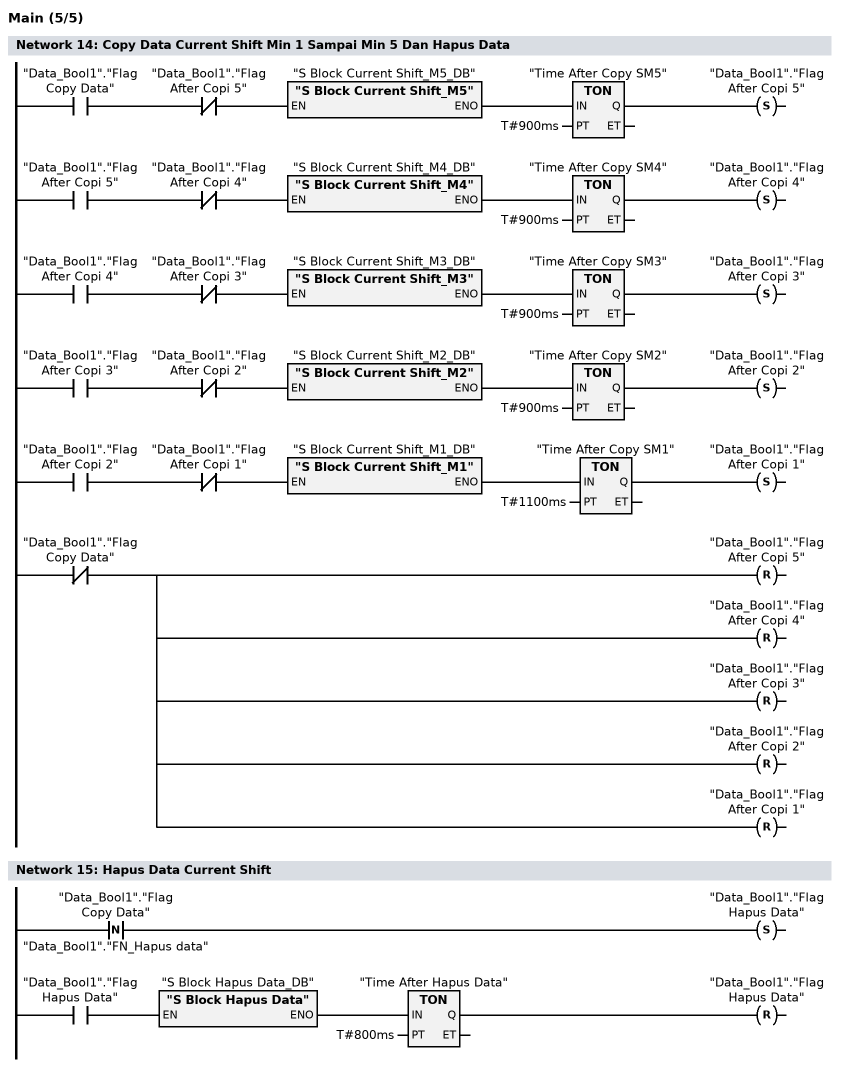
   "S Block Current Shift_M5_DB"(EN := "Data_Bool1"."Flag Copy Data" AND NOT "Data_Bool1"."Flag After Copi 5",   // "S Block Current Shift_M5"
                           ENO => #_w1);
   "Time After Copy SM5".TON(IN := #_w1, PT := T#900ms);
   IF "Time After Copy SM5".Q THEN "Data_Bool1"."Flag After Copi 5" := TRUE; END_IF;
   "S Block Current Shift_M4_DB"(EN := "Data_Bool1"."Flag After Copi 5" AND NOT "Data_Bool1"."Flag After Copi 4",   // "S Block Current Shift_M4"
                           ENO => #_w2);
   "Time After Copy SM4".TON(IN := #_w2, PT := T#900ms);
   IF "Time After Copy SM4".Q THEN "Data_Bool1"."Flag After Copi 4" := TRUE; END_IF;
   "S Block Current Shift_M3_DB"(EN := "Data_Bool1"."Flag After Copi 4" AND NOT "Data_Bool1"."Flag After Copi 3",   // "S Block Current Shift_M3"
                           ENO => #_w3);
   "Time After Copy SM3".TON(IN := #_w3, PT := T#900ms);
   IF "Time After Copy SM3".Q THEN "Data_Bool1"."Flag After Copi 3" := TRUE; END_IF;
   "S Block Current Shift_M2_DB"(EN := "Data_Bool1"."Flag After Copi 3" AND NOT "Data_Bool1"."Flag After Copi 2",   // "S Block Current Shift_M2"
                           ENO => #_w4);
   "Time After Copy SM2".TON(IN := #_w4, PT := T#900ms);
   IF "Time After Copy SM2".Q THEN "Data_Bool1"."Flag After Copi 2" := TRUE; END_IF;
   "S Block Current Shift_M1_DB"(EN := "Data_Bool1"."Flag After Copi 2" AND NOT "Data_Bool1"."Flag After Copi 1",   // "S Block Current Shift_M1"
                           ENO => #_w5);
   "Time After Copy SM1".TON(IN := #_w5, PT := T#1100ms);
   IF "Time After Copy SM1".Q THEN "Data_Bool1"."Flag After Copi 1" := TRUE; END_IF;
   IF NOT "Data_Bool1"."Flag Copy Data" THEN
       "Data_Bool1"."Flag After Copi 5" := FALSE;
       "Data_Bool1"."Flag After Copi 4" := FALSE;
       "Data_Bool1"."Flag After Copi 3" := FALSE;
       "Data_Bool1"."Flag After Copi 2" := FALSE;
       "Data_Bool1"."Flag After Copi 1" := FALSE;
   END_IF;
END_REGION

REGION Network 15: Hapus Data Current Shift
   #_w1 := NOT "Data_Bool1"."Flag Copy Data" AND "Data_Bool1"."FN_Hapus data";   // falling edge of "Data_Bool1"."Flag Copy Data"
   "Data_Bool1"."FN_Hapus data" := "Data_Bool1"."Flag Copy Data";
   IF #_w1 THEN "Data_Bool1"."Flag Hapus Data" := TRUE; END_IF;
   "S Block Hapus Data_DB"(EN := "Data_Bool1"."Flag Hapus Data", ENO => #_w2);   // "S Block Hapus Data"
   "Time After Hapus Data".TON(IN := #_w2, PT := T#800ms);
   IF "Time After Hapus Data".Q THEN "Data_Bool1"."Flag Hapus Data" := FALSE; END_IF;
END_REGION
END_ORGANIZATION_BLOCK

ORGANIZATION_BLOCK "Time error interrupt"   // OB80, LAD, TimeErrorInterrupt
{ S7_Optimized_Access := 'TRUE' }
VERSION : 0.1
   VAR_INPUT
      Fault_ID : Byte;   // Fault identifier
      Csg_OBnr : OB_Any;   // Number of OB causing the error
      Csg_Prio : UInt;   // Priority of OB causing the error
   END_VAR
BEGIN
END_ORGANIZATION_BLOCK

ORGANIZATION_BLOCK "Diagnostic error interrupt"   // OB82, LAD, DiagnosticErrorInterrupt
{ S7_Optimized_Access := 'TRUE' }
VERSION : 0.1
   VAR_INPUT
      IO_State : Word;   // IO state of the HW object
      LADDR : Hw_Any;   // Hardware identifier
      Channel : UInt;   // Channel number
      MultiError : Bool;   // =true if more than one error is present
   END_VAR
BEGIN
END_ORGANIZATION_BLOCK

(* ===== HMI "HMI_RT_1" =====
system functions are stored by id; their names below are inferred from use
connection "HMI_connection": ETHERNET, SMART_S7_1200_OMS

HMI tags "Default tag table"
   "Tag_ScreenNumber" : UInt, internal
      on ChangeValue: ActivateScreenByNumber("Tag_ScreenNumber", 0)
   "PB Test Pneumatic 1" : Bool = PLC "PB Test Pneumatic 1" AT %M205.1, 1 s
   "PB Test Pneumatic 2" : Bool = PLC "PB Test Pneumatic 2" AT %M205.2, 1 s
   "PB Test Pneumatic 3" : Bool = PLC "PB Test Pneumatic 3" AT %M205.3, 1 s
   "PB Test Pneumatic 4" : Bool = PLC "PB Test Pneumatic 4" AT %M205.4, 1 s
   "PB Test Pneumatic 5" : Bool = PLC "PB Test Pneumatic 5" AT %M205.5, 1 s
   "PB Test Motor" : Bool = PLC "PB Test Motor" AT %M205.7, 1 s
   "PB Test Manual Servo" : Bool = PLC "PB Test Manual Servo" AT %M205.6, 1 s
   "Timer Waktu Pemanasan" : Time = PLC "Timer Delay Heating" AT %MD0, 1 s
   "Machine Running" : Bool = PLC "Machine Running" AT %M200.0, 1 s
   "Flag Imaje Start" : Bool = PLC "Flag Imaje Start" AT %M212.0, 1 s
   "Counter" : Int = PLC Counter AT %MW5, 1 s
   "Counter Ejector" : Int = PLC "Counter Ejector" AT %MW9, 1 s
   "Reset Counter" : Bool = PLC "Reset Counter" AT %M200.1, 1 s
   "PB Test Mode" : Bool = PLC "PB Test Mode" AT %M205.0, 1 s
   "Flag Ejector Jalan" : Bool = PLC "Flag Ejector Jalan" AT %M230.3, 1 s
   "Error Group" : Word = PLC "Error Group" AT %MW4, 1 s
   "PB Test Imaje" : Bool = PLC "PB Test Imaje" AT %M206.0, 1 s
   "PB Test Air Valve" : Bool = PLC "PB Test Air Valve" AT %M206.1, 1 s
   "Flag Barcode HMI" : Bool = PLC "Flag Enable/Disable Barcode HMI" AT %M30.0, 1 s
   "Flag Enable/Disable Error Chute 3 Way" : Bool = PLC "Flag Enable/Disable Error Chute 3 Way" AT %M30.1, 1 s
   "Flag Parameter Page" : Bool = PLC "Flag Parameter Page" AT %M232.6, 1 s
   "Flag Main Page" : Bool = PLC "Flag Main Page" AT %M232.7, 1 s
   "HMI_Tag_1" : Word AT %DB39.DBW0, 1 s
   "HMI_Error_Cont" : Word AT %DB40.DBW0, 1 s
   "Flag Teach In Barcode" : Bool = PLC "Flag Teach In Barcode" AT %M212.4, 1 s
   "Teach In Barcode" : Bool = PLC "Teach In Barcode" AT %Q0.5, 1 s
   "Flag Heater Error HMI" : Bool = PLC "Flag Heater Error HMI" AT %M30.2, 1 s
   "Flag Pneumatic Bypass" : Bool = PLC "Flag Reed Switch Bypass" AT %M30.3, 1 s
   "Flag Enable/Disable Error Door Open" : Bool = PLC "Flag Enable/Disable Error Door Open" AT %M30.5, 1 s
   "Timer Delay Stamp" : Time = PLC "Timer Delay Stamp" AT %MD32, 1 s
   "Flag Enable/Disable Block Focke" : Bool = PLC "Flag Enable/Disable Block Focke" AT %M30.6, 1 s
   "Flag Enable/Disable Error Chute Before Heating Roll" : Bool = PLC "Flag Enable/Disable Error Chute Before Heating Roll" AT %M30.4, 1 s
   "Flag Machine Bypass" : Bool = PLC "Flag Machine Bypass" AT %M30.7, 1 s
   "RS Bypass Pneumatic 1" : Bool = PLC "RS Bypass Pneumatic 1" AT %M31.0, 1 s
   "RS Bypass Pneumatic 3" : Bool = PLC "RS Bypass Pneumatic 3" AT %M31.1, 1 s
   "RS Bypass Pneumatic 4" : Bool = PLC "RS Bypass Pneumatic 4" AT %M31.2, 1 s
   "RS Bypass Pneumatic 5" : Bool = PLC "RS Bypass Pneumatic 5" AT %M31.3, 1 s
   "PB Test Pneumatic 6" : Bool = PLC "PB Test Pneumatic 6" AT %M206.2, 1 s
   "PB Test Conveyor" : Bool = PLC "PB Test Conveyor" AT %M206.3, 1 s
   "Flag Enable/Disable Flow to Reject" : Bool = PLC "Flag Enable/Disable Flow to Reject" AT %M31.5, 1 s
   "PB Test Motor Coveyor Pusher" : Bool = PLC "PB Test Motor Coveyor Pusher" AT %M206.4, 1 s
   "PB Test Motor Heating Roll" : Bool = PLC "PB Test Motor Heating Roll" AT %M206.5, 1 s
   "Timer Trigger Barcode" : Time = PLC "Timer Scanning Barcode" AT %MD36, 1 s
   "Flag Enable/Disable Heating Roll" : Bool = PLC "Flag Enable/Disable Heating Roll" AT %M31.6, 1 s
   "Data_DTLData_DTL_Imaje Not In Position[0]" : DTL = PLC Data_DTLData."DTL_Imaje Not In Position"[0], 1 s
   "Data_DTLData_DTL_Imaje Not In Position[0].HOUR" : USInt = PLC Data_DTLData."DTL_Imaje Not In Position"[0].HOUR, 1 s
   "Data_DTLData_DTL_Imaje Not In Position[0].MINUTE" : USInt = PLC Data_DTLData."DTL_Imaje Not In Position"[0].MINUTE, 1 s
   "Data_DTLData_DTL_Imaje Not In Position[0].SECOND" : USInt = PLC Data_DTLData."DTL_Imaje Not In Position"[0].SECOND, 1 s
   "Data_DTLData_DTL_Imaje Not In Position[1].HOUR" : USInt = PLC Data_DTLData."DTL_Imaje Not In Position"[1].HOUR, 1 s
   "Data_DTLData_DTL_Imaje Not In Position[1].MINUTE" : USInt = PLC Data_DTLData."DTL_Imaje Not In Position"[1].MINUTE, 1 s
   "Data_DTLData_DTL_Imaje Not In Position[1].SECOND" : USInt = PLC Data_DTLData."DTL_Imaje Not In Position"[1].SECOND, 1 s
   "Data_DTLData_DTL_Imaje Not In Position[2].HOUR" : USInt = PLC Data_DTLData."DTL_Imaje Not In Position"[2].HOUR, 1 s
   "Data_DTLData_DTL_Imaje Not In Position[2].MINUTE" : USInt = PLC Data_DTLData."DTL_Imaje Not In Position"[2].MINUTE, 1 s
   "Data_DTLData_DTL_Imaje Not In Position[2].SECOND" : USInt = PLC Data_DTLData."DTL_Imaje Not In Position"[2].SECOND, 1 s
   "Data_DTLData_DTL_Imaje Not In Position[3].HOUR" : USInt = PLC Data_DTLData."DTL_Imaje Not In Position"[3].HOUR, 1 s
   "Data_DTLData_DTL_Imaje Not In Position[3].MINUTE" : USInt = PLC Data_DTLData."DTL_Imaje Not In Position"[3].MINUTE, 1 s
   "Data_DTLData_DTL_Imaje Not In Position[3].SECOND" : USInt = PLC Data_DTLData."DTL_Imaje Not In Position"[3].SECOND, 1 s
   "Data_DTLData_DTL_Imaje Not In Position[4].HOUR" : USInt = PLC Data_DTLData."DTL_Imaje Not In Position"[4].HOUR, 1 s
   "Data_DTLData_DTL_Imaje Not In Position[4].MINUTE" : USInt = PLC Data_DTLData."DTL_Imaje Not In Position"[4].MINUTE, 1 s
   "Data_DTLData_DTL_Imaje Not In Position[4].SECOND" : USInt = PLC Data_DTLData."DTL_Imaje Not In Position"[4].SECOND, 1 s
   "Data_DTLData_DTL_Imaje Not In Position[5].HOUR" : USInt = PLC Data_DTLData."DTL_Imaje Not In Position"[5].HOUR, 1 s
   "Data_DTLData_DTL_Imaje Not In Position[5].MINUTE" : USInt = PLC Data_DTLData."DTL_Imaje Not In Position"[5].MINUTE, 1 s
   "Data_DTLData_DTL_Imaje Not In Position[5].SECOND" : USInt = PLC Data_DTLData."DTL_Imaje Not In Position"[5].SECOND, 1 s
   "Data_DTLData_DTL_Mesin Error[0].HOUR" : USInt = PLC Data_DTLData."DTL_Mesin Error"[0].HOUR, 1 s   // Mulai Copi
   "Data_DTLData_DTL_Mesin Error[0].MINUTE" : USInt = PLC Data_DTLData."DTL_Mesin Error"[0].MINUTE, 1 s
   "Data_DTLData_DTL_Mesin Error[0].SECOND" : USInt = PLC Data_DTLData."DTL_Mesin Error"[0].SECOND, 1 s
   "Data_DTLData_DTL_Mesin Error[1].HOUR" : USInt = PLC Data_DTLData."DTL_Mesin Error"[1].HOUR, 1 s
   "Data_DTLData_DTL_Mesin Error[1].MINUTE" : USInt = PLC Data_DTLData."DTL_Mesin Error"[1].MINUTE, 1 s
   "Data_DTLData_DTL_Mesin Error[1].SECOND" : USInt = PLC Data_DTLData."DTL_Mesin Error"[1].SECOND, 1 s
   "Data_DTLData_DTL_Mesin Error[2].HOUR" : USInt = PLC Data_DTLData."DTL_Mesin Error"[2].HOUR, 1 s
   "Data_DTLData_DTL_Mesin Error[2].MINUTE" : USInt = PLC Data_DTLData."DTL_Mesin Error"[2].MINUTE, 1 s
   "Data_DTLData_DTL_Mesin Error[2].SECOND" : USInt = PLC Data_DTLData."DTL_Mesin Error"[2].SECOND, 1 s
   "Data_DTLData_DTL_Mesin Error[3].HOUR" : USInt = PLC Data_DTLData."DTL_Mesin Error"[3].HOUR, 1 s
   "Data_DTLData_DTL_Mesin Error[3].MINUTE" : USInt = PLC Data_DTLData."DTL_Mesin Error"[3].MINUTE, 1 s
   "Data_DTLData_DTL_Mesin Error[3].SECOND" : USInt = PLC Data_DTLData."DTL_Mesin Error"[3].SECOND, 1 s
   "Data_DTLData_DTL_Mesin Error[4].HOUR" : USInt = PLC Data_DTLData."DTL_Mesin Error"[4].HOUR, 1 s
   "Data_DTLData_DTL_Mesin Error[4].MINUTE" : USInt = PLC Data_DTLData."DTL_Mesin Error"[4].MINUTE, 1 s
   "Data_DTLData_DTL_Mesin Error[4].SECOND" : USInt = PLC Data_DTLData."DTL_Mesin Error"[4].SECOND, 1 s
   "Data_DTLData_DTL_Mesin Error[5].HOUR" : USInt = PLC Data_DTLData."DTL_Mesin Error"[5].HOUR, 1 s
   "Data_DTLData_DTL_Mesin Error[5].MINUTE" : USInt = PLC Data_DTLData."DTL_Mesin Error"[5].MINUTE, 1 s
   "Data_DTLData_DTL_Mesin Error[5].SECOND" : USInt = PLC Data_DTLData."DTL_Mesin Error"[5].SECOND, 1 s
   "Data_DTLData_DTL_Mesin Run Baypass[0].HOUR" : USInt = PLC Data_DTLData."DTL_Mesin Run Baypass"[0].HOUR, 1 s
   "Data_DTLData_DTL_Mesin Run Baypass[0].MINUTE" : USInt = PLC Data_DTLData."DTL_Mesin Run Baypass"[0].MINUTE, 1 s
   "Data_DTLData_DTL_Mesin Run Baypass[0].SECOND" : USInt = PLC Data_DTLData."DTL_Mesin Run Baypass"[0].SECOND, 1 s
   "Data_DTLData_DTL_Mesin Run Baypass[1].HOUR" : USInt = PLC Data_DTLData."DTL_Mesin Run Baypass"[1].HOUR, 1 s
   "Data_DTLData_DTL_Mesin Run Baypass[1].MINUTE" : USInt = PLC Data_DTLData."DTL_Mesin Run Baypass"[1].MINUTE, 1 s
   "Data_DTLData_DTL_Mesin Run Baypass[1].SECOND" : USInt = PLC Data_DTLData."DTL_Mesin Run Baypass"[1].SECOND, 1 s
   "Data_DTLData_DTL_Mesin Run Baypass[2].HOUR" : USInt = PLC Data_DTLData."DTL_Mesin Run Baypass"[2].HOUR, 1 s
   "Data_DTLData_DTL_Mesin Run Baypass[2].MINUTE" : USInt = PLC Data_DTLData."DTL_Mesin Run Baypass"[2].MINUTE, 1 s
   "Data_DTLData_DTL_Mesin Run Baypass[2].SECOND" : USInt = PLC Data_DTLData."DTL_Mesin Run Baypass"[2].SECOND, 1 s
   "Data_DTLData_DTL_Mesin Run Baypass[3].HOUR" : USInt = PLC Data_DTLData."DTL_Mesin Run Baypass"[3].HOUR, 1 s
   "Data_DTLData_DTL_Mesin Run Baypass[3].MINUTE" : USInt = PLC Data_DTLData."DTL_Mesin Run Baypass"[3].MINUTE, 1 s
   "Data_DTLData_DTL_Mesin Run Baypass[3].SECOND" : USInt = PLC Data_DTLData."DTL_Mesin Run Baypass"[3].SECOND, 1 s
   "Data_DTLData_DTL_Mesin Run Baypass[4].HOUR" : USInt = PLC Data_DTLData."DTL_Mesin Run Baypass"[4].HOUR, 1 s
   "Data_DTLData_DTL_Mesin Run Baypass[4].MINUTE" : USInt = PLC Data_DTLData."DTL_Mesin Run Baypass"[4].MINUTE, 1 s
   "Data_DTLData_DTL_Mesin Run Baypass[4].SECOND" : USInt = PLC Data_DTLData."DTL_Mesin Run Baypass"[4].SECOND, 1 s
   "Data_DTLData_DTL_Mesin Run Baypass[5].HOUR" : USInt = PLC Data_DTLData."DTL_Mesin Run Baypass"[5].HOUR, 1 s
   "Data_DTLData_DTL_Mesin Run Baypass[5].MINUTE" : USInt = PLC Data_DTLData."DTL_Mesin Run Baypass"[5].MINUTE, 1 s
   "Data_DTLData_DTL_Mesin Run Baypass[5].SECOND" : USInt = PLC Data_DTLData."DTL_Mesin Run Baypass"[5].SECOND, 1 s
   "Data_DTLData_DTL_Mesin Run[0].HOUR" : USInt = PLC Data_DTLData."DTL_Mesin Run"[0].HOUR, 1 s
   "Data_DTLData_DTL_Mesin Run[0].MINUTE" : USInt = PLC Data_DTLData."DTL_Mesin Run"[0].MINUTE, 1 s
   "Data_DTLData_DTL_Mesin Run[0].SECOND" : USInt = PLC Data_DTLData."DTL_Mesin Run"[0].SECOND, 1 s
   "Data_DTLData_DTL_Mesin Run[1].HOUR" : USInt = PLC Data_DTLData."DTL_Mesin Run"[1].HOUR, 1 s
   "Data_DTLData_DTL_Mesin Run[1].MINUTE" : USInt = PLC Data_DTLData."DTL_Mesin Run"[1].MINUTE, 1 s
   "Data_DTLData_DTL_Mesin Run[1].SECOND" : USInt = PLC Data_DTLData."DTL_Mesin Run"[1].SECOND, 1 s
   "Data_DTLData_DTL_Mesin Run[2].HOUR" : USInt = PLC Data_DTLData."DTL_Mesin Run"[2].HOUR, 1 s
   "Data_DTLData_DTL_Mesin Run[2].MINUTE" : USInt = PLC Data_DTLData."DTL_Mesin Run"[2].MINUTE, 1 s
   "Data_DTLData_DTL_Mesin Run[2].SECOND" : USInt = PLC Data_DTLData."DTL_Mesin Run"[2].SECOND, 1 s
   "Data_DTLData_DTL_Mesin Run[3].HOUR" : USInt = PLC Data_DTLData."DTL_Mesin Run"[3].HOUR, 1 s
   "Data_DTLData_DTL_Mesin Run[3].MINUTE" : USInt = PLC Data_DTLData."DTL_Mesin Run"[3].MINUTE, 1 s
   "Data_DTLData_DTL_Mesin Run[3].SECOND" : USInt = PLC Data_DTLData."DTL_Mesin Run"[3].SECOND, 1 s
   "Data_DTLData_DTL_Mesin Run[4].HOUR" : USInt = PLC Data_DTLData."DTL_Mesin Run"[4].HOUR, 1 s
   "Data_DTLData_DTL_Mesin Run[4].MINUTE" : USInt = PLC Data_DTLData."DTL_Mesin Run"[4].MINUTE, 1 s
   "Data_DTLData_DTL_Mesin Run[4].SECOND" : USInt = PLC Data_DTLData."DTL_Mesin Run"[4].SECOND, 1 s
   "Data_DTLData_DTL_Mesin Run[5].HOUR" : USInt = PLC Data_DTLData."DTL_Mesin Run"[5].HOUR, 1 s
   "Data_DTLData_DTL_Mesin Run[5].MINUTE" : USInt = PLC Data_DTLData."DTL_Mesin Run"[5].MINUTE, 1 s
   "Data_DTLData_DTL_Mesin Run[5].SECOND" : USInt = PLC Data_DTLData."DTL_Mesin Run"[5].SECOND, 1 s
   "Data_DTLData_DTL_Mesin Stop[0].HOUR" : USInt = PLC Data_DTLData."DTL_Mesin Stop"[0].HOUR, 1 s
   "Data_DTLData_DTL_Mesin Stop[0].MINUTE" : USInt = PLC Data_DTLData."DTL_Mesin Stop"[0].MINUTE, 1 s
   "Data_DTLData_DTL_Mesin Stop[0].SECOND" : USInt = PLC Data_DTLData."DTL_Mesin Stop"[0].SECOND, 1 s
   "Data_DTLData_DTL_Mesin Stop[1].HOUR" : USInt = PLC Data_DTLData."DTL_Mesin Stop"[1].HOUR, 1 s
   "Data_DTLData_DTL_Mesin Stop[1].MINUTE" : USInt = PLC Data_DTLData."DTL_Mesin Stop"[1].MINUTE, 1 s
   "Data_DTLData_DTL_Mesin Stop[1].SECOND" : USInt = PLC Data_DTLData."DTL_Mesin Stop"[1].SECOND, 1 s
   "Data_DTLData_DTL_Mesin Stop[2].HOUR" : USInt = PLC Data_DTLData."DTL_Mesin Stop"[2].HOUR, 1 s
   "Data_DTLData_DTL_Mesin Stop[2].MINUTE" : USInt = PLC Data_DTLData."DTL_Mesin Stop"[2].MINUTE, 1 s
   "Data_DTLData_DTL_Mesin Stop[2].SECOND" : USInt = PLC Data_DTLData."DTL_Mesin Stop"[2].SECOND, 1 s
   "Data_DTLData_DTL_Mesin Stop[3].HOUR" : USInt = PLC Data_DTLData."DTL_Mesin Stop"[3].HOUR, 1 s
   "Data_DTLData_DTL_Mesin Stop[3].MINUTE" : USInt = PLC Data_DTLData."DTL_Mesin Stop"[3].MINUTE, 1 s
   "Data_DTLData_DTL_Mesin Stop[3].SECOND" : USInt = PLC Data_DTLData."DTL_Mesin Stop"[3].SECOND, 1 s
   "Data_DTLData_DTL_Mesin Stop[4].HOUR" : USInt = PLC Data_DTLData."DTL_Mesin Stop"[4].HOUR, 1 s
   "Data_DTLData_DTL_Mesin Stop[4].MINUTE" : USInt = PLC Data_DTLData."DTL_Mesin Stop"[4].MINUTE, 1 s
   "Data_DTLData_DTL_Mesin Stop[4].SECOND" : USInt = PLC Data_DTLData."DTL_Mesin Stop"[4].SECOND, 1 s
   "Data_DTLData_DTL_Mesin Stop[5].HOUR" : USInt = PLC Data_DTLData."DTL_Mesin Stop"[5].HOUR, 1 s
   "Data_DTLData_DTL_Mesin Stop[5].MINUTE" : USInt = PLC Data_DTLData."DTL_Mesin Stop"[5].MINUTE, 1 s
   "Data_DTLData_DTL_Mesin Stop[5].SECOND" : USInt = PLC Data_DTLData."DTL_Mesin Stop"[5].SECOND, 1 s   // akhir copi
   "Data_DTLData_DTL_Paper R Out[0].HOUR" : USInt = PLC Data_DTLData."DTL_Paper R Out"[0].HOUR, 1 s
   "Data_DTLData_DTL_Paper R Out[0].MINUTE" : USInt = PLC Data_DTLData."DTL_Paper R Out"[0].MINUTE, 1 s
   "Data_DTLData_DTL_Paper R Out[0].SECOND" : USInt = PLC Data_DTLData."DTL_Paper R Out"[0].SECOND, 1 s
   "Data_DTLData_DTL_Paper R Out[1].HOUR" : USInt = PLC Data_DTLData."DTL_Paper R Out"[1].HOUR, 1 s
   "Data_DTLData_DTL_Paper R Out[1].MINUTE" : USInt = PLC Data_DTLData."DTL_Paper R Out"[1].MINUTE, 1 s
   "Data_DTLData_DTL_Paper R Out[1].SECOND" : USInt = PLC Data_DTLData."DTL_Paper R Out"[1].SECOND, 1 s
   "Data_DTLData_DTL_Paper R Out[2].HOUR" : USInt = PLC Data_DTLData."DTL_Paper R Out"[2].HOUR, 1 s
   "Data_DTLData_DTL_Paper R Out[2].MINUTE" : USInt = PLC Data_DTLData."DTL_Paper R Out"[2].MINUTE, 1 s
   "Data_DTLData_DTL_Paper R Out[2].SECOND" : USInt = PLC Data_DTLData."DTL_Paper R Out"[2].SECOND, 1 s
   "Data_DTLData_DTL_Paper R Out[3].HOUR" : USInt = PLC Data_DTLData."DTL_Paper R Out"[3].HOUR, 1 s
   "Data_DTLData_DTL_Paper R Out[3].MINUTE" : USInt = PLC Data_DTLData."DTL_Paper R Out"[3].MINUTE, 1 s
   "Data_DTLData_DTL_Paper R Out[3].SECOND" : USInt = PLC Data_DTLData."DTL_Paper R Out"[3].SECOND, 1 s
   "Data_DTLData_DTL_Paper R Out[4].HOUR" : USInt = PLC Data_DTLData."DTL_Paper R Out"[4].HOUR, 1 s
   "Data_DTLData_DTL_Paper R Out[4].MINUTE" : USInt = PLC Data_DTLData."DTL_Paper R Out"[4].MINUTE, 1 s
   "Data_DTLData_DTL_Paper R Out[5].HOUR" : USInt = PLC Data_DTLData."DTL_Paper R Out"[5].HOUR, 1 s
   "Data_DTLData_DTL_Paper R Out[5].MINUTE" : USInt = PLC Data_DTLData."DTL_Paper R Out"[5].MINUTE, 1 s
   "Data_DTLData_DTL_Paper R Out[5].SECOND" : USInt = PLC Data_DTLData."DTL_Paper R Out"[5].SECOND, 1 s
   "Data_IntData_Frekuensi Error[1]" : USInt = PLC Data_IntData."Frekuensi Error"[1], 1 s
   "Data_IntData_Frekuensi Error[2]" : USInt = PLC Data_IntData."Frekuensi Error"[2], 1 s
   "Data_IntData_Frekuensi Error[3]" : USInt = PLC Data_IntData."Frekuensi Error"[3], 1 s
   "Data_IntData_Frekuensi Error[4]" : USInt = PLC Data_IntData."Frekuensi Error"[4], 1 s
   "Data_IntData_Frekuensi Error[5]" : USInt = PLC Data_IntData."Frekuensi Error"[5], 1 s
   "Data_IntData_Frekuensi Error[6]" : USInt = PLC Data_IntData."Frekuensi Error"[6], 1 s
   "Data_IntData_Frekuensi Error[7]" : USInt = PLC Data_IntData."Frekuensi Error"[7], 1 s
   "Data_IntData_Frekuensi Error_1[1]" : USInt = PLC Data_IntData."Frekuensi Error_1"[1], 1 s
   "Data_IntData_Frekuensi Error_1[2]" : USInt = PLC Data_IntData."Frekuensi Error_1"[2], 1 s
   "Data_IntData_Frekuensi Error_1[3]" : USInt = PLC Data_IntData."Frekuensi Error_1"[3], 1 s
   "Data_IntData_Frekuensi Error_1[4]" : USInt = PLC Data_IntData."Frekuensi Error_1"[4], 1 s
   "Data_IntData_Frekuensi Error_1[5]" : USInt = PLC Data_IntData."Frekuensi Error_1"[5], 1 s
   "Data_IntData_Frekuensi Error_1[6]" : USInt = PLC Data_IntData."Frekuensi Error_1"[6], 1 s
   "Data_IntData_Frekuensi Error_1[7]" : USInt = PLC Data_IntData."Frekuensi Error_1"[7], 1 s
   "Data_IntData_Frekuensi Error_2[1]" : USInt = PLC Data_IntData."Frekuensi Error_2"[1], 1 s
   "Data_IntData_Frekuensi Error_2[2]" : USInt = PLC Data_IntData."Frekuensi Error_2"[2], 1 s
   "Data_IntData_Frekuensi Error_2[3]" : USInt = PLC Data_IntData."Frekuensi Error_2"[3], 1 s
   "Data_IntData_Frekuensi Error_2[4]" : USInt = PLC Data_IntData."Frekuensi Error_2"[4], 1 s
   "Data_IntData_Frekuensi Error_2[5]" : USInt = PLC Data_IntData."Frekuensi Error_2"[5], 1 s
   "Data_IntData_Frekuensi Error_2[6]" : USInt = PLC Data_IntData."Frekuensi Error_2"[6], 1 s
   "Data_IntData_Frekuensi Error_2[7]" : USInt = PLC Data_IntData."Frekuensi Error_2"[7], 1 s
   "Data_IntData_Frekuensi Error_3[1]" : USInt = PLC Data_IntData."Frekuensi Error_3"[1], 1 s
   "Data_IntData_Frekuensi Error_3[2]" : USInt = PLC Data_IntData."Frekuensi Error_3"[2], 1 s
   "Data_IntData_Frekuensi Error_3[3]" : USInt = PLC Data_IntData."Frekuensi Error_3"[3], 1 s
   "Data_IntData_Frekuensi Error_3[4]" : USInt = PLC Data_IntData."Frekuensi Error_3"[4], 1 s
   "Data_IntData_Frekuensi Error_3[5]" : USInt = PLC Data_IntData."Frekuensi Error_3"[5], 1 s
   "Data_IntData_Frekuensi Error_3[6]" : USInt = PLC Data_IntData."Frekuensi Error_3"[6], 1 s
   "Data_IntData_Frekuensi Error_3[7]" : USInt = PLC Data_IntData."Frekuensi Error_3"[7], 1 s
   "Data_IntData_Frekuensi Error_4[1]" : USInt = PLC Data_IntData."Frekuensi Error_4"[1], 1 s
   "Data_IntData_Frekuensi Error_4[2]" : USInt = PLC Data_IntData."Frekuensi Error_4"[2], 1 s
   "Data_IntData_Frekuensi Error_4[3]" : USInt = PLC Data_IntData."Frekuensi Error_4"[3], 1 s
   "Data_IntData_Frekuensi Error_4[4]" : USInt = PLC Data_IntData."Frekuensi Error_4"[4], 1 s
   "Data_IntData_Frekuensi Error_4[5]" : USInt = PLC Data_IntData."Frekuensi Error_4"[5], 1 s
   "Data_IntData_Frekuensi Error_4[6]" : USInt = PLC Data_IntData."Frekuensi Error_4"[6], 1 s
   "Data_IntData_Frekuensi Error_4[7]" : USInt = PLC Data_IntData."Frekuensi Error_4"[7], 1 s
   "Data_IntData_Frekuensi Error_5[1]" : USInt = PLC Data_IntData."Frekuensi Error_5"[1], 1 s
   "Data_IntData_Frekuensi Error_5[2]" : USInt = PLC Data_IntData."Frekuensi Error_5"[2], 1 s
   "Data_IntData_Frekuensi Error_5[3]" : USInt = PLC Data_IntData."Frekuensi Error_5"[3], 1 s
   "Data_IntData_Frekuensi Error_5[4]" : USInt = PLC Data_IntData."Frekuensi Error_5"[4], 1 s
   "Data_IntData_Frekuensi Error_5[5]" : USInt = PLC Data_IntData."Frekuensi Error_5"[5], 1 s
   "Data_IntData_Frekuensi Error_5[6]" : USInt = PLC Data_IntData."Frekuensi Error_5"[6], 1 s
   "Data_IntData_Frekuensi Error_5[7]" : USInt = PLC Data_IntData."Frekuensi Error_5"[7], 1 s
   "Data_integer2_Flag Input Always bad Read" : USInt = PLC Data_integer2."Flag Input Always bad Read", 1 s
   "Data_Real_% Total Output[0]" : Real = PLC Data_Real."% Total Output"[0], 1 s
   "Data_Real_% Total Output[1]" : Real = PLC Data_Real."% Total Output"[1], 1 s
   "Data_Real_% Total Output[2]" : Real = PLC Data_Real."% Total Output"[2], 1 s
   "Data_Real_% Total Output[3]" : Real = PLC Data_Real."% Total Output"[3], 1 s
   "Data_Real_% Total Output[4]" : Real = PLC Data_Real."% Total Output"[4], 1 s
   "Data_Real_% Total Output[5]" : Real = PLC Data_Real."% Total Output"[5], 1 s
   "Data_Real_%Downstream stop[0]" : Real = PLC Data_Real."%Downstream stop"[0], 1 s
   "Data_Real_%Mesin Error[0]" : Real = PLC Data_Real."%Mesin Error"[0], 1 s   // Mulai copi 2
   "Data_Real_%Mesin Error[1]" : Real = PLC Data_Real."%Mesin Error"[1], 1 s
   "Data_Real_%Mesin Error[2]" : Real = PLC Data_Real."%Mesin Error"[2], 1 s
   "Data_Real_%Mesin Error[3]" : Real = PLC Data_Real."%Mesin Error"[3], 1 s
   "Data_Real_%Mesin Error[4]" : Real = PLC Data_Real."%Mesin Error"[4], 1 s
   "Data_Real_%Mesin Error[5]" : Real = PLC Data_Real."%Mesin Error"[5], 1 s
   "Data_Real_%Mesin Run Baypass[0]" : Real = PLC Data_Real."%Mesin Run Baypass"[0], 1 s
   "Data_Real_%Mesin Run Baypass[1]" : Real = PLC Data_Real."%Mesin Run Baypass"[1], 1 s
   "Data_Real_%Mesin Run Baypass[2]" : Real = PLC Data_Real."%Mesin Run Baypass"[2], 1 s
   "Data_Real_%Mesin Run Baypass[3]" : Real = PLC Data_Real."%Mesin Run Baypass"[3], 1 s
   "Data_Real_%Mesin Run Baypass[4]" : Real = PLC Data_Real."%Mesin Run Baypass"[4], 1 s
   "Data_Real_%Mesin Run Baypass[5]" : Real = PLC Data_Real."%Mesin Run Baypass"[5], 1 s
   "Data_Real_%Mesin Run[0]" : Real = PLC Data_Real."%Mesin Run"[0], 1 s
   "Data_Real_%Mesin Run[1]" : Real = PLC Data_Real."%Mesin Run"[1], 1 s
   "Data_Real_%Mesin Run[2]" : Real = PLC Data_Real."%Mesin Run"[2], 1 s
   "Data_Real_%Mesin Run[3]" : Real = PLC Data_Real."%Mesin Run"[3], 1 s
   "Data_Real_%Mesin Run[4]" : Real = PLC Data_Real."%Mesin Run"[4], 1 s
   "Data_Real_%Mesin Run[5]" : Real = PLC Data_Real."%Mesin Run"[5], 1 s
   "Data_Real_%Mesin Stop[0]" : Real = PLC Data_Real."%Mesin Stop"[0], 1 s
   "Data_Real_%Mesin Stop[1]" : Real = PLC Data_Real."%Mesin Stop"[1], 1 s
   "Data_Real_%Mesin Stop[2]" : Real = PLC Data_Real."%Mesin Stop"[2], 1 s
   "Data_Real_%Mesin Stop[3]" : Real = PLC Data_Real."%Mesin Stop"[3], 1 s
   "Data_Real_%Mesin Stop[4]" : Real = PLC Data_Real."%Mesin Stop"[4], 1 s
   "Data_Real_%Mesin Stop[5]" : Real = PLC Data_Real."%Mesin Stop"[5], 1 s   // Stop Copi 2
   "DB_Bool1_F_Set Time Day" : Bool = PLC Data_Bool1."F_Set Time Day", 1 s
   "DB_Bool1_F_Set Time Shift" : Bool = PLC Data_Bool1."F_Set Time Shift", 1 s
   "DB_DTL1_Cur_ShiftA" : DTL = PLC Data_DTL1.Cur_ShiftA, 1 s
   "DB_DTL1_Cur_ShiftA_1" : DTL = PLC Data_DTL1.Cur_ShiftA_1, 1 s
   "DB_DTL1_Cur_ShiftA_2" : DTL = PLC Data_DTL1.Cur_ShiftA_2, 1 s
   "DB_DTL1_Cur_ShiftA_3" : DTL = PLC Data_DTL1.Cur_ShiftA_3, 1 s
   "DB_DTL1_Cur_ShiftA_4" : DTL = PLC Data_DTL1.Cur_ShiftA_4, 1 s
   "DB_DTL1_Cur_ShiftA_5" : DTL = PLC Data_DTL1.Cur_ShiftA_5, 1 s
   "DB_DTL1_Cur_ShiftB" : DTL = PLC Data_DTL1.Cur_ShiftB, 1 s
   "DB_DTL1_Cur_ShiftB_1" : DTL = PLC Data_DTL1.Cur_ShiftB_1, 1 s
   "DB_DTL1_Cur_ShiftB_2" : DTL = PLC Data_DTL1.Cur_ShiftB_2, 1 s
   "DB_DTL1_Cur_ShiftB_3" : DTL = PLC Data_DTL1.Cur_ShiftB_3, 1 s
   "DB_DTL1_Cur_ShiftB_4" : DTL = PLC Data_DTL1.Cur_ShiftB_4, 1 s
   "DB_DTL1_Cur_ShiftB_5" : DTL = PLC Data_DTL1.Cur_ShiftB_5, 1 s
   "DB_DTL1_Input" : DTL = PLC Data_DTL1.Input, 1 s
   "DB_DTL1_Input.DAY" : USInt = PLC Data_DTL1.Input.DAY, 1 s
   "DB_DTL1_Output" : DTL = PLC Data_DTL1.Output, 1 s
   "DB_DTLData_DTL_Down Stop.HOUR" : USInt = PLC Data_DTLData."DTL_Down Stop".HOUR, 1 s
   "DB_DTLData_DTL_Down Stop.MINUTE" : USInt = PLC Data_DTLData."DTL_Down Stop".MINUTE, 1 s
   "DB_DTLData_DTL_Down Stop.SECOND" : USInt = PLC Data_DTLData."DTL_Down Stop".SECOND, 1 s
   "DB_DTLData_DTL_Down Stop_1.HOUR" : USInt = PLC Data_DTLData."DTL_Down Stop_1".HOUR, 1 s
   "DB_DTLData_DTL_Down Stop_1.MINUTE" : USInt = PLC Data_DTLData."DTL_Down Stop_1".MINUTE, 1 s
   "DB_DTLData_DTL_Down Stop_1.SECOND" : USInt = PLC Data_DTLData."DTL_Down Stop_1".SECOND, 1 s
   "DB_DTLData_DTL_Down Stop_2.HOUR" : USInt = PLC Data_DTLData."DTL_Down Stop_2".HOUR, 1 s
   "DB_DTLData_DTL_Down Stop_2.MINUTE" : USInt = PLC Data_DTLData."DTL_Down Stop_2".MINUTE, 1 s
   "DB_DTLData_DTL_Down Stop_2.SECOND" : USInt = PLC Data_DTLData."DTL_Down Stop_2".SECOND, 1 s
   "DB_DTLData_DTL_Down Stop_3.HOUR" : USInt = PLC Data_DTLData."DTL_Down Stop_3".HOUR, 1 s
   "DB_DTLData_DTL_Down Stop_3.MINUTE" : USInt = PLC Data_DTLData."DTL_Down Stop_3".MINUTE, 1 s
   "DB_DTLData_DTL_Down Stop_3.SECOND" : USInt = PLC Data_DTLData."DTL_Down Stop_3".SECOND, 1 s
   "DB_DTLData_DTL_Down Stop_4.HOUR" : USInt = PLC Data_DTLData."DTL_Down Stop_4".HOUR, 1 s
   "DB_DTLData_DTL_Down Stop_4.MINUTE" : USInt = PLC Data_DTLData."DTL_Down Stop_4".MINUTE, 1 s
   "DB_DTLData_DTL_Down Stop_4.SECOND" : USInt = PLC Data_DTLData."DTL_Down Stop_4".SECOND, 1 s
   "DB_DTLData_DTL_Down Stop_5.HOUR" : USInt = PLC Data_DTLData."DTL_Down Stop_5".HOUR, 1 s
   "DB_DTLData_DTL_Down Stop_5.MINUTE" : USInt = PLC Data_DTLData."DTL_Down Stop_5".MINUTE, 1 s
   "DB_DTLData_DTL_Down Stop_5.SECOND" : USInt = PLC Data_DTLData."DTL_Down Stop_5".SECOND, 1 s
   "DB_DTLData_DTL_Imaje Er.HOUR" : USInt = PLC Data_DTLData."DTL_Imaje Er".HOUR, 1 s
   "DB_DTLData_DTL_Imaje Er.MINUTE" : USInt = PLC Data_DTLData."DTL_Imaje Er".MINUTE, 1 s
   "DB_DTLData_DTL_Imaje Er.SECOND" : USInt = PLC Data_DTLData."DTL_Imaje Er".SECOND, 1 s
   "DB_DTLData_DTL_Imaje Er_1.HOUR" : USInt = PLC Data_DTLData."DTL_Imaje Er_1".HOUR, 1 s
   "DB_DTLData_DTL_Imaje Er_1.MINUTE" : USInt = PLC Data_DTLData."DTL_Imaje Er_1".MINUTE, 1 s
   "DB_DTLData_DTL_Imaje Er_1.SECOND" : USInt = PLC Data_DTLData."DTL_Imaje Er_1".SECOND, 1 s
   "DB_DTLData_DTL_Imaje Er_2.HOUR" : USInt = PLC Data_DTLData."DTL_Imaje Er_2".HOUR, 1 s
   "DB_DTLData_DTL_Imaje Er_2.MINUTE" : USInt = PLC Data_DTLData."DTL_Imaje Er_2".MINUTE, 1 s
   "DB_DTLData_DTL_Imaje Er_2.SECOND" : USInt = PLC Data_DTLData."DTL_Imaje Er_2".SECOND, 1 s
   "DB_DTLData_DTL_Imaje Er_3.HOUR" : USInt = PLC Data_DTLData."DTL_Imaje Er_3".HOUR, 1 s
   "DB_DTLData_DTL_Imaje Er_3.MINUTE" : USInt = PLC Data_DTLData."DTL_Imaje Er_3".MINUTE, 1 s
   "DB_DTLData_DTL_Imaje Er_3.SECOND" : USInt = PLC Data_DTLData."DTL_Imaje Er_3".SECOND, 1 s
   "DB_DTLData_DTL_Imaje Er_4.HOUR" : USInt = PLC Data_DTLData."DTL_Imaje Er_4".HOUR, 1 s
   "DB_DTLData_DTL_Imaje Er_4.MINUTE" : USInt = PLC Data_DTLData."DTL_Imaje Er_4".MINUTE, 1 s
   "DB_DTLData_DTL_Imaje Er_4.SECOND" : USInt = PLC Data_DTLData."DTL_Imaje Er_4".SECOND, 1 s
   "DB_DTLData_DTL_Imaje Er_5.HOUR" : USInt = PLC Data_DTLData."DTL_Imaje Er_5".HOUR, 1 s
   "DB_DTLData_DTL_Imaje Er_5.MINUTE" : USInt = PLC Data_DTLData."DTL_Imaje Er_5".MINUTE, 1 s
   "DB_DTLData_DTL_Imaje Er_5.SECOND" : USInt = PLC Data_DTLData."DTL_Imaje Er_5".SECOND, 1 s
   "DB_DTLData_DTL_Press Low.HOUR" : USInt = PLC Data_DTLData."DTL_Press Low".HOUR, 1 s
   "DB_DTLData_DTL_Press Low.MINUTE" : USInt = PLC Data_DTLData."DTL_Press Low".MINUTE, 1 s
   "DB_DTLData_DTL_Press Low.SECOND" : USInt = PLC Data_DTLData."DTL_Press Low".SECOND, 1 s
   "DB_DTLData_DTL_Press Low_1.HOUR" : USInt = PLC Data_DTLData."DTL_Press Low_1".HOUR, 1 s
   "DB_DTLData_DTL_Press Low_1.MINUTE" : USInt = PLC Data_DTLData."DTL_Press Low_1".MINUTE, 1 s
   "DB_DTLData_DTL_Press Low_1.SECOND" : USInt = PLC Data_DTLData."DTL_Press Low_1".SECOND, 1 s
   "DB_DTLData_DTL_Press Low_2.HOUR" : USInt = PLC Data_DTLData."DTL_Press Low_2".HOUR, 1 s
   "DB_DTLData_DTL_Press Low_2.MINUTE" : USInt = PLC Data_DTLData."DTL_Press Low_2".MINUTE, 1 s
   "DB_DTLData_DTL_Press Low_2.SECOND" : USInt = PLC Data_DTLData."DTL_Press Low_2".SECOND, 1 s
   "DB_DTLData_DTL_Press Low_3.HOUR" : USInt = PLC Data_DTLData."DTL_Press Low_3".HOUR, 1 s
   "DB_DTLData_DTL_Press Low_3.MINUTE" : USInt = PLC Data_DTLData."DTL_Press Low_3".MINUTE, 1 s
   "DB_DTLData_DTL_Press Low_3.SECOND" : USInt = PLC Data_DTLData."DTL_Press Low_3".SECOND, 1 s
   "DB_DTLData_DTL_Press Low_4.HOUR" : USInt = PLC Data_DTLData."DTL_Press Low_4".HOUR, 1 s
   "DB_DTLData_DTL_Press Low_4.MINUTE" : USInt = PLC Data_DTLData."DTL_Press Low_4".MINUTE, 1 s
   "DB_DTLData_DTL_Press Low_4.SECOND" : USInt = PLC Data_DTLData."DTL_Press Low_4".SECOND, 1 s
   "DB_DTLData_DTL_Press Low_5.HOUR" : USInt = PLC Data_DTLData."DTL_Press Low_5".HOUR, 1 s
   "DB_DTLData_DTL_Press Low_5.MINUTE" : USInt = PLC Data_DTLData."DTL_Press Low_5".MINUTE, 1 s
   "DB_DTLData_DTL_Press Low_5.SECOND" : USInt = PLC Data_DTLData."DTL_Press Low_5".SECOND, 1 s
   "DB_DTLData_DTL_RS Pneu Er.HOUR" : USInt = PLC Data_DTLData."DTL_RS Pneu Er".HOUR, 1 s
   "DB_DTLData_DTL_RS Pneu Er.MINUTE" : USInt = PLC Data_DTLData."DTL_RS Pneu Er".MINUTE, 1 s
   "DB_DTLData_DTL_RS Pneu Er.SECOND" : USInt = PLC Data_DTLData."DTL_RS Pneu Er".SECOND, 1 s
   "DB_DTLData_DTL_RS Pneu Er_1.HOUR" : USInt = PLC Data_DTLData."DTL_RS Pneu Er_1".HOUR, 1 s
   "DB_DTLData_DTL_RS Pneu Er_1.MINUTE" : USInt = PLC Data_DTLData."DTL_RS Pneu Er_1".MINUTE, 1 s
   "DB_DTLData_DTL_RS Pneu Er_1.SECOND" : USInt = PLC Data_DTLData."DTL_RS Pneu Er_1".SECOND, 1 s
   "DB_DTLData_DTL_RS Pneu Er_2.HOUR" : USInt = PLC Data_DTLData."DTL_RS Pneu Er_2".HOUR, 1 s
   "DB_DTLData_DTL_RS Pneu Er_2.MINUTE" : USInt = PLC Data_DTLData."DTL_RS Pneu Er_2".MINUTE, 1 s
   "DB_DTLData_DTL_RS Pneu Er_2.SECOND" : USInt = PLC Data_DTLData."DTL_RS Pneu Er_2".SECOND, 1 s
   "DB_DTLData_DTL_RS Pneu Er_3.HOUR" : USInt = PLC Data_DTLData."DTL_RS Pneu Er_3".HOUR, 1 s
   "DB_DTLData_DTL_RS Pneu Er_3.MINUTE" : USInt = PLC Data_DTLData."DTL_RS Pneu Er_3".MINUTE, 1 s
   "DB_DTLData_DTL_RS Pneu Er_3.SECOND" : USInt = PLC Data_DTLData."DTL_RS Pneu Er_3".SECOND, 1 s
   "DB_DTLData_DTL_RS Pneu Er_4.HOUR" : USInt = PLC Data_DTLData."DTL_RS Pneu Er_4".HOUR, 1 s
   "DB_DTLData_DTL_RS Pneu Er_4.MINUTE" : USInt = PLC Data_DTLData."DTL_RS Pneu Er_4".MINUTE, 1 s
   "DB_DTLData_DTL_RS Pneu Er_4.SECOND" : USInt = PLC Data_DTLData."DTL_RS Pneu Er_4".SECOND, 1 s
   "DB_DTLData_DTL_RS Pneu Er_5.HOUR" : USInt = PLC Data_DTLData."DTL_RS Pneu Er_5".HOUR, 1 s
   "DB_DTLData_DTL_RS Pneu Er_5.MINUTE" : USInt = PLC Data_DTLData."DTL_RS Pneu Er_5".MINUTE, 1 s
   "DB_DTLData_DTL_RS Pneu Er_5.SECOND" : USInt = PLC Data_DTLData."DTL_RS Pneu Er_5".SECOND, 1 s
   "DB_DTLData_DTL_Slof Jam.HOUR" : USInt = PLC Data_DTLData."DTL_Slof Jam".HOUR, 1 s
   "DB_DTLData_DTL_Slof Jam.MINUTE" : USInt = PLC Data_DTLData."DTL_Slof Jam".MINUTE, 1 s
   "DB_DTLData_DTL_Slof Jam.SECOND" : USInt = PLC Data_DTLData."DTL_Slof Jam".SECOND, 1 s
   "DB_DTLData_DTL_Slof Jam_1.HOUR" : USInt = PLC Data_DTLData."DTL_Slof Jam_1".HOUR, 1 s
   "DB_DTLData_DTL_Slof Jam_1.MINUTE" : USInt = PLC Data_DTLData."DTL_Slof Jam_1".MINUTE, 1 s
   "DB_DTLData_DTL_Slof Jam_1.SECOND" : USInt = PLC Data_DTLData."DTL_Slof Jam_1".SECOND, 1 s
   "DB_DTLData_DTL_Slof Jam_2.HOUR" : USInt = PLC Data_DTLData."DTL_Slof Jam_2".HOUR, 1 s
   "DB_DTLData_DTL_Slof Jam_2.MINUTE" : USInt = PLC Data_DTLData."DTL_Slof Jam_2".MINUTE, 1 s
   "DB_DTLData_DTL_Slof Jam_2.SECOND" : USInt = PLC Data_DTLData."DTL_Slof Jam_2".SECOND, 1 s
   "DB_DTLData_DTL_Slof Jam_3.HOUR" : USInt = PLC Data_DTLData."DTL_Slof Jam_3".HOUR, 1 s
   "DB_DTLData_DTL_Slof Jam_3.MINUTE" : USInt = PLC Data_DTLData."DTL_Slof Jam_3".MINUTE, 1 s
   "DB_DTLData_DTL_Slof Jam_3.SECOND" : USInt = PLC Data_DTLData."DTL_Slof Jam_3".SECOND, 1 s
   "DB_DTLData_DTL_Slof Jam_4.HOUR" : USInt = PLC Data_DTLData."DTL_Slof Jam_4".HOUR, 1 s
   "DB_DTLData_DTL_Slof Jam_4.MINUTE" : USInt = PLC Data_DTLData."DTL_Slof Jam_4".MINUTE, 1 s
   "DB_DTLData_DTL_Slof Jam_4.SECOND" : USInt = PLC Data_DTLData."DTL_Slof Jam_4".SECOND, 1 s
   "DB_DTLData_DTL_Slof Jam_5.HOUR" : USInt = PLC Data_DTLData."DTL_Slof Jam_5".HOUR, 1 s
   "DB_DTLData_DTL_Slof Jam_5.MINUTE" : USInt = PLC Data_DTLData."DTL_Slof Jam_5".MINUTE, 1 s
   "DB_DTLData_DTL_Slof Jam_5.SECOND" : USInt = PLC Data_DTLData."DTL_Slof Jam_5".SECOND, 1 s
   "DB_IntData_Bad R" : UDInt = PLC Data_IntData."Bad R", 1 s
   "DB_IntData_Bad R_1" : UDInt = PLC Data_IntData."Bad R_1", 1 s
   "DB_IntData_Bad R_2" : UDInt = PLC Data_IntData."Bad R_2", 1 s
   "DB_IntData_Bad R_3" : UDInt = PLC Data_IntData."Bad R_3", 1 s
   "DB_IntData_Bad R_4" : UDInt = PLC Data_IntData."Bad R_4", 1 s
   "DB_IntData_Bad R_5" : UDInt = PLC Data_IntData."Bad R_5", 1 s
   "DB_IntData_Good R1" : UDInt = PLC Data_IntData."Good R", 1 s
   "DB_IntData_Good R1_1" : UDInt = PLC Data_IntData."Good R_1", 1 s
   "DB_IntData_Good R1_2" : UDInt = PLC Data_IntData."Good R_2", 1 s
   "DB_IntData_Good R1_3" : UDInt = PLC Data_IntData."Good R_3", 1 s
   "DB_IntData_Good R1_4" : UDInt = PLC Data_IntData."Good R_4", 1 s
   "DB_IntData_Good R1_5" : UDInt = PLC Data_IntData."Good R_5", 1 s
   "DB_IntData_Good R2" : UDInt = PLC Data_IntData."Reject Out S", 1 s
   "DB_IntData_Good R2_1" : UDInt = PLC Data_IntData."Reject Out S_1", 1 s
   "DB_IntData_Good R2_2" : UDInt = PLC Data_IntData."Reject Out S_2", 1 s
   "DB_IntData_Good R2_3" : UDInt = PLC Data_IntData."Reject Out S_3", 1 s
   "DB_IntData_Good R2_4" : UDInt = PLC Data_IntData."Reject Out S_4", 1 s
   "DB_IntData_Good R2_5" : UDInt = PLC Data_IntData."Reject Out S_5", 1 s
   "DB_IntData_Input Sloft" : UDInt = PLC Data_IntData."Input Sloft", 1 s
   "DB_IntData_Input Sloft_1" : UDInt = PLC Data_IntData."Input Sloft_1", 1 s
   "DB_IntData_Input Sloft_2" : UDInt = PLC Data_IntData."Input Sloft_2", 1 s
   "DB_IntData_Input Sloft_3" : UDInt = PLC Data_IntData."Input Sloft_3", 1 s
   "DB_IntData_Input Sloft_4" : UDInt = PLC Data_IntData."Input Sloft_4", 1 s
   "DB_IntData_Input Sloft_5" : UDInt = PLC Data_IntData."Input Sloft_5", 1 s
   "DB_IntData_Tot Good R" : UDInt = PLC Data_IntData."Tot Out Slof", 1 s
   "DB_IntData_Tot Good R_2" : UDInt = PLC Data_IntData."Tot Out Slof_2", 1 s
   "DB_IntData_Tot Good R_3" : UDInt = PLC Data_IntData."Tot Out Slof_3", 1 s
   "DB_IntData_Tot Good R_4" : UDInt = PLC Data_IntData."Tot Out Slof_4", 1 s
   "DB_IntData_Tot Good R_5" : UDInt = PLC Data_IntData."Tot Out Slof_5", 1 s
   "DB_IntData_Tot Out Slof_1" : UDInt = PLC Data_IntData."Tot Out Slof_1", 1 s
   "DB_Integer_IDay" : USInt = PLC Data_Integer.IDay, 1 s